screen "Screen_Doseerwals" 800x480, template "Popup_Parameters_Manual"
   on GenerateScreen: SetBit("HMI_ManualControl")
   on ClearScreen: ResetBit("HMI_ManualControl")
   TextField "Text field_1" at 624,181 size 48x23; Text 'Ready'
      Visibility <- "Drive 3 Ready"
   TextField "Text field_5" at 628,181 size 74x23; Text 'Not ready'
      Visibility <- "Drive 3 Ready"
   TextField "Template_Text field_1" at 423,141 size 182x23; Text 'Walzen - Parameters'
   TextField "Text field_3" at 10,228 size 192x23; Text 'Handbediening Walzen'
   TextField "Text field_8" at 85,262 size 42x23; Text 'Rust'
      Visibility <- "Drive 3 RUN FWD"
   TextField "Text field_9" at 103,262 size 111x23; Text 'Wals running'
      Visibility <- "Drive 3 RUN FWD"
   TextField "Text field_4" at 433,180 size 105x23; Text 'Drive Status'
   TextField "Text field_6" at 433,354 size 165x23; Text 'Reference Position:'
   IOField "StartMotorTimer" at 626,350 size 96x32; FormatPattern 9999
      ProcessValue <- "PositionManagement_Axis 3_Values_Reference Position"
   TextField "Text field_12" at 433,395 size 113x23; Text 'Rest Position'
   IOField "I/O field_2" at 625,392 size 96x32; FormatPattern 99.9999
      ProcessValue <- "PositionManagement_Axis 3_Values_Rest Position"
   Button "Button_5" at 16,389 size 111x66; TextOff '++'
      Appearance <- "Drive_3_Manual"
      on Press: SetBit("Manual Jog Fwd")
      on Release: ResetBit("Manual Jog Fwd")
   Button "Button_6" at 152,388 size 111x66; TextOff '--'
      on Release: ResetBit("Manual Jog Rev")
      on Press: SetBit("Manual Jog Rev")
   Circle "Circle_1" at 626,206 size 20x20
      Appearance <- "Voorverdeelwals staat in positie"
   Group "Group_DriveStatus" at 624,181 size 78x23
   GraphicView "Graphic view_1" at 210,135 size 172x116; Picture "MotoriconArrowLeftRight"
   Circle "Circle_2" at 221,181 size 20x20
      Appearance <- "Drive 3 REV"
   Circle "Circle_3" at 344,181 size 20x20
      Appearance <- "Drive 3 RUN FWD"
   Circle "Circle_4" at 264,229 size 16x16
      Appearance <- "Drive 3 Rapid Stop"
   TextField "Text field_2" at 210,225 size 53x23; Text 'Brake'
   TextField "Text field_10" at 13,314 size 144x23; Text 'Current Position:'
   IOField "I/O field_1" at 160,307 size 140x35; FormatPattern 9999.9999
      ProcessValue <- "PositionManagement_Data_Actual_Axis1_Position"
   TextField "Text field_11" at 433,206 size 148x23; Text 'Reference Sensor'
   TextField "Text field_13" at 433,235 size 163x23; Text 'Pulsfactor Encoder:'
   IOField "I/O field_3" at 626,229 size 96x32; FormatPattern 999.99
      ProcessValue <- "PositionManagement_Axis 3_Values_Pulsfactor"
   TextField "Text field_14" at 13,347 size 144x23; Text 'Desired Position:'
   IOField "I/O field_4" at 160,343 size 140x35; FormatPattern 999.9
      ProcessValue <- "PositionManagement_Demo_Pos_Desired_Pos"
   Button "Button_7" at 314,348 size 45x26; TextOff 'Go'
      on Press: SetBit("PositionManagement_Demo_Pos_Start")
      on Release: ResetBit("PositionManagement_Demo_Pos_Start")
   TextField "Text field_15" at 313,310 size 59x22; Text 'Degrees'
   TextField "Text field_16" at 434,275 size 101x23; Text 'Axis Speed:'
   IOField "I/O field_5" at 626,269 size 96x32; FormatPattern 99
      ProcessValue <- "PositionManagement_Axis 3_Values_Axis_Speed"
   TextField "Text field_17" at 434,314 size 163x23; Text 'Position Tolerance:'
   IOField "I/O field_6" at 626,308 size 96x32; FormatPattern 9.99
      ProcessValue <- "PositionManagement_Axis 3_Values_Position Offset"
   TextField "Text field_18" at 726,354 size 59x22; Text 'Degrees'
   TextField "Text field_19" at 727,315 size 59x22; Text 'Degrees'
   TextField "Text field_20" at 729,274 size 20x22; Text '%'
   TextField "Text field_21" at 731,234 size 41x22; Text 'Steps'
   TextField "Text field_22" at 728,396 size 59x22; Text 'Degrees'
   TextField "Text field_7" at 433,431 size 92x23; Text 'Raw Value'
   IOField "I/O field_7" at 625,428 size 96x32; FormatPattern 999999
      ProcessValue <- "Counter2_IW102"
   TextField "Text field_23" at 728,432 size 45x22; Text 'Pulses'
   Button "Button_1" at 16,149 size 126x32; TextOff 'Start Ref Run'
      on Release: ResetBit("PositionManagement_Axis 3_Commands_Start Ref Run")
      on Press: SetBit("PositionManagement_Axis 3_Commands_Start Ref Run")
      Appearance <- "Drive_3_Manual"

screen "Screen_Afdichting" 800x480, template "Popup_Parameters_Manual"
   on GenerateScreen: SetBit("HMI_ManualControl")
   on ClearScreen: ResetBit("HMI_ManualControl")
   TextField "Text field_2" at 10,228 size 290x23; Text 'Handbediening Afdichtingssysteem'
   TextField "Text field_8" at 85,262 size 42x23; Text 'Rust'
      Visibility <- "Valve 1"
   TextField "Text field_9" at 103,262 size 120x23; Text 'Valve opening'
      Visibility <- "Valve 1"
   TextField "Text field_6" at 477,376 size 247x23; Text 'Currently no parameters here'
   TextField "Template_Text field_1" at 430,142 size 205x23; Text 'Afdichting - Parameters'
   TextField "Template_Text field_2" at 12,307 size 232x23; Text 'Afdichting - Handbediening'
   Button "Button_1" at 25,340 size 110x70; TextOff 'Cilinder uit'
      on Click: SetBit("Valve_1_Manual")
      Appearance <- "Valve_1_Manual"
   Button "Button_2" at 152,340 size 110x70; TextOff 'Cilinder in'
      on Click: ResetBit("Valve_1_Manual")
   Group "Enable_Module_2" at 278,358 size 99x32; TextList "Enable / Disable List"; PictureList "Enable_Graphic"
   Group "Group" at 533,189 size 143x74; Picture "Pneumatic 5_2 valve"
   GraphicView "Graphic view_1" at 533,199 size 143x64; Picture "Pneumatic 5_2 valve"
   Circle "Circle_1" at 536,189 size 20x20
      Appearance <- "Valve 1"
   SymbolicIOField "Symbolic I/O field_3" at 311,358 size 66x32; TextOn '1'; TextOff '0'; TextList "Enable / Disable List"
      ProcessValue <- "PLCMemory_Disable_Modules_Disable_Afsluiter"
   GraphicIOField "Graphic I/O field_3" at 278,358 size 32x32; PictureList "Enable_Graphic"
      on Deactivate: ResetBit("PLCMemory_Disable_Modules_Disable_Aandruk1")
      on Activate: SetBit("PLCMemory_Disable_Modules_Disable_Aandruk1")
      ProcessValue <- "PLCMemory_Disable_Modules_Disable_Afsluiter"

screen "Screen_Settings" 800x480, template "Popup_Parameters_Manual"
   TextField "Text field_1" at 7,129 size 141x23; Text 'General Settings'
   Button "Button_7" at 487,6 size 96x65; TextOff 'Home'
      on Click: ActivateScreen("Screen_Handbediening", 0)
   TextField "Text field_12" at 420,218 size 131x23; Text 'Wals Slip Time:'
   IOField "Wals_Slip_Time" at 656,213 size 96x32; FormatPattern 9999
      ProcessValue <- "PLCMemory_WalsCheck_Time"
   TextField "Text field_13" at 420,255 size 174x23; Text 'Magazijn leeg delay:'
   IOField "I/O field_2" at 656,251 size 96x32; FormatPattern 99999
      ProcessValue <- "PLCMemory_Magazijn_Sensor_Delay"
   TextField "Template_Text field_1" at 420,154 size 186x23; Text 'General - Parameters'
   Button "Button_5" at 16,189 size 333x55; TextOff 'Manual Start'
      on Click: SetBit("RUN_Manual")
   Button "Button_6" at 15,255 size 333x55; TextOff 'Manual Stop'
      on Click: ResetBit("RUN_Manual")
   TextField "Text field_3" at 11,156 size 371x23; Text 'DO NOT USE THIS BUTTONS! IT IS DANGEROUS!'
   IOField "I/O field_1" at 656,173 size 96x32; FormatPattern 9999
      ProcessValue <- "PLCMemory_Safety_Delay"
   TextField "Text field_2" at 421,177 size 137x23; Text 'Safety on delay:'
   Button "Button_9" at 23,420 size 122x32; TextOff 'Close RT'
      on Click: StopRuntime(0)
   Button "Button_10" at 156,420 size 122x32; TextOff 'Alarms / LOG'
      on Click: ActivateScreen("AlarmWindow", 0)
   TextField "Text field_4" at 16,325 size 118x23; Text 'Invert Safety:'
   TextField "Text field_5" at 16,362 size 168x23; Text 'Invert Notensensor:'
   SymbolicIOField "Symbolic I/O field_1" at 253,317 size 96x32; TextOff '0'; TextOn '1'; TextList "List_Deactivate_Module"
      ProcessValue <- "Safety_Override"
   SymbolicIOField "Symbolic I/O field_2" at 253,353 size 96x32; TextOn '1'; TextOff '0'; TextList "List_Deactivate_Module"
      ProcessValue <- "Invert_Trechter_Sensor"
   TextField "Text field_8" at 420,295 size 174x23; Text 'Product Check Time:'
   IOField "ProductCheckTime" at 656,291 size 96x32; FormatPattern 99999
      ProcessValue <- "PLCMemory_ProductCheck_Time"
   IOField "I/O field_3" at 658,403 size 96x32; FormatPattern 999999
      ProcessValue <- "PLCMemory_TD_Products_Counter"
   TextField "Text field_6" at 422,407 size 229x23; Text 'Aantal producten gedraaid:'
   Button "Button_11" at 659,440 size 122x32; TextOff 'Reset teller'
      on Press: SetBit("ResetTotalProducts")
      on Release: ResetBit("ResetTotalProducts")
   TextField "Text field_11" at 754,176 size 25x22; Text 'ms'
   TextField "Text field_7" at 754,216 size 25x22; Text 'ms'
   TextField "Text field_9" at 754,253 size 25x22; Text 'ms'
   TextField "Text field_10" at 754,293 size 25x22; Text 'ms'
   TextField "Text field_14" at 421,334 size 169x23; Text 'BlowOff Cycle Time:'
   IOField "ProductCheckTime_1" at 657,330 size 96x32; FormatPattern 99999
      ProcessValue <- "PLCMemory_Offset_Timers_BlowOff_CycleTime"
   TextField "Text field_15" at 755,332 size 25x22; Text 'ms'
   TextField "Text field_16" at 422,372 size 170x23; Text 'BlowOff Pulse Time:'
   IOField "ProductCheckTime_2" at 658,367 size 96x32; FormatPattern 99999
      ProcessValue <- "PLCMemory_Offset_Timers_Blow_Off_PulseTime"
   TextField "Text field_17" at 756,369 size 25x22; Text 'ms'
   Softkey "Softkey_F1" at 0,0 size 0x0
      on KeyDown: function_ee5b8808("Button_7")
      on KeyUp: function_f101fd67("Button_7")

Template "Popup_Parameters" 800x480
   Rectangle "Rectangle_1" at 0,33 size 799x45
      Visibility <- "Alarm_Product_Not_Position"
   TextField "Text field_2" at 99,41 size 644x29; Text 'Aanvoer - Producten komen niet op positie, controleer sensor'
      Visibility <- "Alarm_Product_Not_Position"
   GraphicView "Graphic view_1" at 8,39 size 37x35; Picture "Graphic_30"
      Visibility <- "Alarm_Product_Not_Position"
   Group "ProductNotPositionError_1" at 0,33 size 799x45; Picture "Graphic_30"
   Group "WalsNotPositionError_1" at 0,23 size 799x45; Picture "Graphic_30"
   Group "MagazineEmptyError_1" at 0,11 size 799x45; Picture "Graphic_30"
   Group "ESB_Active_Message_2" at 0,4 size 799x45; Picture "Graphic_31"
   Group "ESB_Active_Message_1" at 1,0 size 799x45; Picture "Graphic_31"
   Rectangle "Rectangle_2" at 0,23 size 799x45
      Visibility <- "Alarm_Axis_Not_Position"
   TextField "Text field_3" at 196,31 size 395x29; Text 'Wals - As komt niet op positie of slipt'
      Visibility <- "Alarm_Axis_Not_Position"
   GraphicView "Graphic view_2" at 8,29 size 37x35; Picture "Graphic_30"
      Visibility <- "Alarm_Axis_Not_Position"
   Rectangle "Rectangle_7" at 0,11 size 799x45
      Visibility <- "Trechter_Bijvullen_Signaal"
   TextField "Text field_4" at 53,19 size 705x29; Text 'Notenmagazijn leeg - Let op, noten bijvullen om te kunnen starten!'
      Visibility <- "Trechter_Bijvullen_Signaal"
   GraphicView "Graphic view_8" at 8,17 size 37x35; Picture "Graphic_30"
      Visibility <- "Trechter_Bijvullen_Signaal"
   Rectangle "Rectangle_8" at 1,0 size 799x45
      Visibility <- "ESB_Safety_Alarm"
   GraphicView "Graphic view_9" at 10,6 size 37x35; Picture "Graphic_31"
      Visibility <- "ESB_Safety_Alarm"
   TextField "Text field_5" at 80,8 size 648x29; Text 'NOODSTOP INGEDRUKT - Ontgrendel Noodstop en druk reset'
      Visibility <- "ESB_Safety_Alarm"
   GraphicView "Graphic view_10" at 753,7 size 37x35; Picture "Graphic_31"
      Visibility <- "ESB_Safety_Alarm"
   Rectangle "Rectangle_3" at 0,4 size 799x45
      Visibility <- "Door_Safety_Alarm"
   GraphicView "Graphic view_3" at 9,10 size 37x35; Picture "Graphic_31"
      Visibility <- "Door_Safety_Alarm"
   TextField "Text field_1" at 174,12 size 511x29; Text 'DEUR(EN) OPEN - Sluit alle deuren en druk reset'
      Visibility <- "Door_Safety_Alarm"
   GraphicView "Graphic view_4" at 752,11 size 37x35; Picture "Graphic_31"
      Visibility <- "Door_Safety_Alarm"
   Group "Message_Group_General" at 0,0 size 800x78; Picture "Graphic_30"

Template "Popup_Parameters_Manual" 800x480
   Rectangle "Rectangle_1" at 0,106 size 799x45
      Visibility <- "Alarm_Product_Not_Position"
   TextField "Text field_2" at 99,114 size 644x29; Text 'Aanvoer - Producten komen niet op positie, controleer sensor'
      Visibility <- "Alarm_Product_Not_Position"
   GraphicView "Graphic view_1" at 8,112 size 37x35; Picture "Graphic_30"
      Visibility <- "Alarm_Product_Not_Position"
   Group "ProductNotPositionError_1" at 0,106 size 799x45; Picture "Graphic_30"
   Group "WalsNotPositionError_1" at 0,96 size 799x45; Picture "Graphic_30"
   Group "MagazineEmptyError_1" at 0,84 size 799x45; Picture "Graphic_30"
   Group "ESB_Active_Message_2" at 0,77 size 799x45; Picture "Graphic_31"
   Group "ESB_Active_Message_1" at 1,73 size 799x45; Picture "Graphic_31"
   Rectangle "Rectangle_2" at 0,96 size 799x45
      Visibility <- "Alarm_Axis_Not_Position"
   TextField "Text field_3" at 196,104 size 395x29; Text 'Wals - As komt niet op positie of slipt'
      Visibility <- "Alarm_Axis_Not_Position"
   GraphicView "Graphic view_2" at 8,102 size 37x35; Picture "Graphic_30"
      Visibility <- "Alarm_Axis_Not_Position"
   Rectangle "Rectangle_7" at 0,84 size 799x45
      Visibility <- "Trechter_Bijvullen_Signaal"
   TextField "Text field_4" at 53,92 size 705x29; Text 'Notenmagazijn leeg - Let op, noten bijvullen om te kunnen starten!'
      Visibility <- "Trechter_Bijvullen_Signaal"
   GraphicView "Graphic view_8" at 8,90 size 37x35; Picture "Graphic_30"
      Visibility <- "Trechter_Bijvullen_Signaal"
   Rectangle "Rectangle_3" at 0,77 size 799x45
      Visibility <- "Door_Safety_Alarm"
   GraphicView "Graphic view_3" at 9,83 size 37x35; Picture "Graphic_31"
      Visibility <- "Door_Safety_Alarm"
   TextField "Text field_1" at 174,85 size 511x29; Text 'DEUR(EN) OPEN - Sluit alle deuren en druk reset'
      Visibility <- "Door_Safety_Alarm"
   GraphicView "Graphic view_4" at 752,84 size 37x35; Picture "Graphic_31"
      Visibility <- "Door_Safety_Alarm"
   Rectangle "Rectangle_8" at 1,73 size 799x45
      Visibility <- "ESB_Safety_Alarm"
   GraphicView "Graphic view_9" at 10,79 size 37x35; Picture "Graphic_31"
      Visibility <- "ESB_Safety_Alarm"
   TextField "Text field_5" at 80,81 size 648x29; Text 'NOODSTOP INGEDRUKT - Ontgrendel Noodstop en druk reset'
      Visibility <- "ESB_Safety_Alarm"
   GraphicView "Graphic view_10" at 753,80 size 37x35; Picture "Graphic_31"
      Visibility <- "ESB_Safety_Alarm"
   TextField "Text field_7" at 14,261 size 70x23; Text 'Sturing:'
   Button "Button_3" at 693,5 size 100x65; TextOff 'Logoff'
      on Click: function_f23ef4c9()
   Button "Button_4" at 585,5 size 100x65; TextOff 'Back'
      on Click: function_efd93a16()
   Group "Message_Group_Manual" at 0,73 size 800x78; Picture "Graphic_30"

screen "Screen_Automatiek" 800x480, template "Popup_Parameters"
   Softkey "Softkey_F8" at 0,0 size 0x0
      on KeyDown: function_ee5b8808("Button_3")
      on KeyUp: function_f101fd67("Button_3")
   TextField "Text field_1" at 263,165 size 182x23; Text 'Gekozen Programma:'
   TextField "Text field_2" at 451,166 size 15x23; Text '1'
      Appearance <- "LED Programma 1"
   TextField "Text field_3" at 469,166 size 15x23; Text '2'
      Appearance <- "LED Programma 2"
   TextField "Text field_4" at 489,166 size 15x23; Text '3'
      Appearance <- "LED Programma 3"
   Button "Button_3" at 6,157 size 130x60; TextOn 'Onderweg na vorig scherm'; TextOff 'Terug'
      on Click: function_efd93a16()
   Button "Button_1" at 6,222 size 130x60; TextOn 'Onderweg na vorig scherm'; TextOff 'Instellingen'
      on Click: ActivateScreen("Screen_Settings", 0)
   TextField "Text field_5" at 26,112 size 106x23; Text 'Automatiek'
   TextField "Text field_6" at 608,165 size 144x23; Text 'Product Interval:'
   IOField "I/O field_1" at 610,189 size 96x32; FormatPattern 99999
      ProcessValue <- "PLCMemory_ProductIntervalTime"
   TextField "Text field_11" at 710,197 size 68x22; Text 'Seconden'
   TextField "Text field_7" at 292,263 size 179x23; Text 'Aanvoerband Gestart'
      Appearance <- "Drive 1 Ready"
      Visibility <- "Drive 1 RUN FWD"
   TextField "Text field_8" at 299,224 size 160x23; Text 'Koek gedetecteerd'
      Visibility <- "Sensor_op_band_memory"
   TextField "Text field_9" at 290,374 size 178x23; Text 'Doseerwals Draaiend'
      Appearance <- "Drive 3 Ready"
      Visibility <- "PLCMemory_ProductBuffer_MoveTrigger"
   TextField "Text field_10" at 282,337 size 196x23; Text 'Aanvoer Wals Draaiend'
      Visibility <- "Drive 4 RUN FWD"
   TextField "Text field_12" at 308,300 size 146x23; Text 'Trilgoten Gestart'
      Appearance <- "Drive 2 Ready"
      Visibility <- "Drive 2 RUN FWD"
   TextField "Text field_13" at 306,189 size 166x23; Text 'Programma Started'
      Visibility <- "Systeem RUN"
   TextField "Text field_14" at 308,419 size 155x23; Text 'Programma Ended'
      Visibility <- "Systeem RUN"
   GraphicView "Graphic view_1" at 371,209 size 26x22; Picture "Graphic_32"
   GraphicView "Graphic view_2" at 371,246 size 26x22; Picture "Graphic_32"
   GraphicView "Graphic view_3" at 372,283 size 26x22; Picture "Graphic_32"
   GraphicView "Graphic view_4" at 371,320 size 26x22; Picture "Graphic_32"
   GraphicView "Graphic view_5" at 372,357 size 26x22; Picture "Graphic_32"
   GraphicView "Graphic view_6" at 372,399 size 26x22; Picture "Graphic_32"
   TextField "Text field_15" at 608,222 size 123x23; Text 'Product Buffer'
   IOField "I/O field_2" at 610,246 size 96x32; FormatPattern 999
      ProcessValue <- "PLCMemory_ProductBuffer_ProductsCount"
   TextField "Text field_16" at 710,254 size 70x22; Text 'Producten'
   TextField "Text field_17" at 608,281 size 129x23; Text 'Aandruk Buffer'
   IOField "I/O field_3" at 610,305 size 96x32; FormatPattern 99
      ProcessValue <- "PLCMemory_ProductBufferBehindWals_Product_Count"
   TextField "Text field_18" at 710,313 size 70x22; Text 'Producten'
   Button "Button_2" at 6,286 size 130x60; TextOn 'Onderweg na vorig scherm'; TextOff 'Buffer Data'
      on Click: ActivateScreen("Screen_Automatiek_BufferData", 0)

screen "Screen_Trechterwissel" 800x480, template "Popup_Parameters_Manual"
   TextField "Text field_2" at 10,228 size 324x23; Text 'Handbediening Trechter wisselsysteem'
   TextField "Text field_8" at 85,262 size 42x23; Text 'Rust'
      Visibility <- "Valve 2"
   TextField "Text field_9" at 103,262 size 120x23; Text 'Valve opening'
      Visibility <- "Valve 2"
   TextField "Template_Text field_1" at 423,142 size 241x23; Text 'Wisselsysteem - Parameters'
   TextField "Template_Text field_2" at 12,307 size 268x23; Text 'Wisselsysteem - Handbediening'
   Button "Button_1" at 17,338 size 111x32; TextOff 'Cilinder uit'
      on Click: SetBit("Valve_2_Manual")
      Appearance <- "Valve_2_Manual"
   Button "Button_2" at 152,338 size 111x32; TextOff 'Cilinder in'
      on Click: ResetBit("Valve_2_Manual")
   GraphicView "Graphic view_1" at 533,197 size 143x64; Picture "Pneumatic 5_2 valve"
   Circle "Circle_1" at 536,187 size 20x20
      Appearance <- "Valve 2"
   TextField "Text field_13" at 12,381 size 173x23; Text 'Reedcontact Cilinder in:'
   Circle "Circle_2" at 198,384 size 20x20
      Appearance <- "Cilinder Trechterwissel in"
   TextField "Text field_1" at 12,407 size 178x23; Text 'Reedcontact Cilinder uit:'
   Circle "Circle_3" at 198,410 size 20x20
      Appearance <- "Cilinder Trechterwissel uit"
   TextField "Text field_12" at 429,337 size 181x23; Text 'Delay Wisselsysteem:'
   IOField "I/O field_2" at 620,334 size 96x32; FormatPattern 9999

screen "Screen_Aandrukken" 800x480, template "Popup_Parameters_Manual"
   on ClearScreen: ResetBit("HMI_ManualControl")
   on GenerateScreen: SetBit("HMI_ManualControl")
   TextField "Text field_2" at 10,228 size 268x23; Text 'Handbediening Aandruksysteem'
   TextField "Text field_8" at 85,262 size 42x23; Text 'Rust'
      Visibility <- "Valve 3"
   TextField "Text field_9" at 103,262 size 120x23; Text 'Valve opening'
      Visibility <- "Valve 3"
   Button "Button_1" at 428,144 size 110x70; TextOff 'Cilinder 1 uit'
      on Click: SetBit("Valve_3_Manual")
      Appearance <- "Valve_3_Manual"
   Button "Button_2" at 555,144 size 110x70; TextOff 'Cilinder 1 in'
      on Click: ResetBit("Valve_3_Manual")
   Button "Button_5" at 428,241 size 110x70; TextOff 'Cilinder 2 uit'
      on Click: SetBit("Valve_4_Manual")
      Appearance <- "Valve_4_Manual"
   Button "Button_6" at 555,241 size 110x70; TextOff 'Cilinder 2 in'
      on Click: ResetBit("Valve_4_Manual")
   Button "Button_7" at 428,338 size 110x70; TextOff 'Cilinder 3 uit'
      on Click: SetBit("Valve_5_Manual")
      Appearance <- "Valve_5_Manual"
   Button "Button_8" at 555,338 size 110x70; TextOff 'Cilinder 3 in'
      on Click: ResetBit("Valve_5_Manual")
   Button "Button_10" at 24,402 size 150x55; TextOff 'Alle cilinders uit'
      on Click: SetBit("Valve_3_Manual"); SetBit("Valve_4_Manual"); SetBit("Valve_5_Manual")
      Appearance <- "Valve_3_Manual"
   Button "Button_11" at 218,402 size 150x55; TextOff 'Alle cilinders in'
      on Click: ResetBit("Valve_3_Manual"); ResetBit("Valve_4_Manual"); ResetBit("Valve_5_Manual")
   Group "Group" at 15,301 size 207x87; Picture "Pneumatic 5_2 valve"
   Button "Button_3" at 127,351 size 150x45; TextOff 'Blaaspuls aan'
      Appearance <- "Valve_3_Manual"
      on Release: ResetBit("Valve_2_Manual")
      on Press: SetBit("Valve_2_Manual")
   Group "Enable_Module" at 684,163 size 99x32; TextList "Enable / Disable List"; PictureList "Enable_Graphic"
   Group "Enable_Module_1" at 683,264 size 99x32; TextList "Enable / Disable List"; PictureList "Enable_Graphic"
   Group "Enable_Module_2" at 684,357 size 99x32; PictureList "Enable_Graphic"; TextList "Enable / Disable List"
   Group "Enable_Module_3" at 279,356 size 99x32; TextList "Enable / Disable List"; PictureList "Enable_Graphic"
   GraphicView "Graphic view_1" at 16,307 size 95x37; Picture "Pneumatic 5_2 valve"
   GraphicView "Graphic view_2" at 127,307 size 95x37; Picture "Pneumatic 5_2 valve"
   Circle "Circle_2" at 130,301 size 12x12
      Appearance <- "Valve 5"
   Circle "Circle_1" at 19,301 size 12x12
      Appearance <- "Valve 3"
   GraphicView "Graphic view_3" at 15,351 size 95x37; Picture "Pneumatic 5_2 valve"
   Circle "Circle_3" at 18,345 size 12x12
      Appearance <- "Valve 4"
   TextField "Text field_1" at 64,304 size 15x23; Text '1'
   TextField "Text field_3" at 64,348 size 15x23; Text '2'
   TextField "Text field_4" at 176,305 size 15x23; Text '3'
   SymbolicIOField "Symbolic I/O field_2" at 717,163 size 66x32; TextOn '1'; TextOff '0'; TextList "Enable / Disable List"
      ProcessValue <- "PLCMemory_Disable_Modules_Disable_Aandruk1"
   GraphicIOField "Graphic I/O field_1" at 684,163 size 32x32; PictureList "Enable_Graphic"
      ProcessValue <- "PLCMemory_Disable_Modules_Disable_Aandruk1"
      on Activate: SetBit("PLCMemory_Disable_Modules_Disable_Aandruk1")
      on Deactivate: ResetBit("PLCMemory_Disable_Modules_Disable_Aandruk1")
   SymbolicIOField "Symbolic I/O field_1" at 716,264 size 66x32; TextOn '1'; TextOff '0'; TextList "Enable / Disable List"
      ProcessValue <- "PLCMemory_Disable_Modules_Disable_Aandruk2"
   GraphicIOField "Graphic I/O field_2" at 683,264 size 32x32; PictureList "Enable_Graphic"
      on Deactivate: ResetBit("PLCMemory_Disable_Modules_Disable_Aandruk1")
      on Activate: SetBit("PLCMemory_Disable_Modules_Disable_Aandruk1")
      ProcessValue <- "PLCMemory_Disable_Modules_Disable_Aandruk2"
   SymbolicIOField "Symbolic I/O field_3" at 717,357 size 66x32; TextOn '1'; TextOff '0'; TextList "Enable / Disable List"
      ProcessValue <- "PLCMemory_Disable_Modules_Disable_Aandruk3"
   GraphicIOField "Graphic I/O field_3" at 684,357 size 32x32; PictureList "Enable_Graphic"
      on Deactivate: ResetBit("PLCMemory_Disable_Modules_Disable_Aandruk1")
      on Activate: SetBit("PLCMemory_Disable_Modules_Disable_Aandruk1")
      ProcessValue <- "PLCMemory_Disable_Modules_Disable_Aandruk3"
   SymbolicIOField "Symbolic I/O field_4" at 312,356 size 66x32; TextOn '1'; TextOff '0'; TextList "Enable / Disable List"
      ProcessValue <- "PLCMemory_Disable_Modules_Disable_Blaaspuls"
   GraphicIOField "Graphic I/O field_4" at 279,356 size 32x32; PictureList "Enable_Graphic"
      on Deactivate: ResetBit("PLCMemory_Disable_Modules_Disable_Aandruk1")
      on Activate: SetBit("PLCMemory_Disable_Modules_Disable_Aandruk1")
      ProcessValue <- "PLCMemory_Disable_Modules_Disable_Blaaspuls"

screen "Screen_RetourBand" 800x480, template "Popup_Parameters_Manual"
   on GenerateScreen: SetBit("HMI_ManualControl")
   on ClearScreen: ResetBit("HMI_ManualControl")
   TextField "Text field_1" at 8,220 size 255x23; Text 'Handbediening Retoursysteem'
   TextField "Text field_8" at 85,261 size 42x23; Text 'Rust'
      Visibility <- "Drive 5 Ready"
   TextField "Text field_9" at 103,261 size 113x23; Text 'Band running'
      Visibility <- "Drive 5 Ready"
   TextField "Text field_3" at 426,174 size 105x23; Text 'Drive Status'
   TextField "Text field_2" at 426,228 size 153x23; Text 'Start Timer motor'
   IOField "StartMotorTimer" at 584,224 size 96x32; FormatPattern 9999
   TextField "Text field_6" at 426,262 size 149x23; Text 'Stop Timer motor'
   IOField "I/O field_2" at 584,259 size 96x32; FormatPattern 9999
   TextField "Template_Text field_1" at 426,140 size 218x23; Text 'Retourband - Parameters'
   Button "Button_1" at 25,306 size 135x70; TextOff 'Start FWD'
      on Click: SetBit("Drive_5_Manual")
      Appearance <- "Drive_1_Manual"
   Button "Button_2" at 205,306 size 135x70; TextOff 'Stop FWD'
      on Click: ResetBit("Drive_5_Manual")
      on Release: ResetBit("Stop_drive_1")
      on Press: SetBit("Stop_drive_1")
   Button "Button_5" at 25,390 size 135x70; TextOff 'Start Rev'
      on Click: SetBit("Drive 5 REV")
      Appearance <- "Drive 5 REV"
   Button "Button_6" at 205,390 size 135x70; TextOff 'Stop Rev'
      on Click: ResetBit("Drive 5 REV")
   Group "Group" at 582,174 size 77x23
   GraphicView "Graphic view_1" at 272,133 size 135x113; Picture "MotoriconArrowLeftRight"
   Circle "Circle_1" at 277,176 size 20x20
      Appearance <- "Drive 5 REV"
   Circle "Circle_2" at 377,176 size 20x20
      Appearance <- "Drive 5 RUN FWD"
   Circle "Circle_3" at 585,199 size 20x20
      Appearance <- "Drive 5 Rapid Stop"
   TextField "Text field_12" at 426,200 size 101x23; Text 'Drive Brake'
   TextField "Text field_13" at 688,228 size 25x22; Text 'ms'
   TextField "Text field_14" at 688,265 size 25x22; Text 'ms'
   Group "Enable_Module" at 584,298 size 96x32; TextList "Enable / Disable List"; PictureList "Enable_Graphic"
   TextField "Text field_7" at 426,302 size 108x23; Text 'Enable Drive'
   TextField "Text field_5" at 582,174 size 48x23; Text 'Ready'
      Visibility <- "Drive 5 Ready"
   TextField "Text field_4" at 585,174 size 74x23; Text 'Not ready'
      Visibility <- "Drive 5 Ready"
   SymbolicIOField "Symbolic I/O field_2" at 616,298 size 64x32; TextOn '1'; TextOff '0'; TextList "Enable / Disable List"
      ProcessValue <- "PLCMemory_Disable_Modules_Disable_Retourband"
   GraphicIOField "Graphic I/O field_1" at 584,298 size 31x32; PictureList "Enable_Graphic"
      on Deactivate: ResetBit("PLCMemory_Disable_Modules_Disable_Aandruk1")
      on Activate: SetBit("PLCMemory_Disable_Modules_Disable_Aandruk1")
      ProcessValue <- "PLCMemory_Disable_Modules_Disable_Retourband"

screen "Screen_Safety_I/O" 800x480, template "Popup_Parameters"
   TextField "Text field_1" at 185,162 size 145x23; Text 'Noodstop Status:'
   Button "Button_4" at 6,157 size 130x60; TextOn 'Onderweg na vorig scherm'; TextOff 'Terug'
      on Click: function_efd93a16()
   Button "Button_5" at 6,221 size 130x60; TextOn 'Onderweg na vorig scherm'; TextOff 'Instellingen'
      on Click: ActivateScreen("Screen_Settings", 0)
   TextField "Text field_2" at 26,112 size 173x23; Text 'Safety In en Outputs'
   TextField "Text field_6" at 185,221 size 122x23; Text 'Deur 1 Status:'
   TextField "Text field_3" at 185,252 size 122x23; Text 'Deur 2 Status:'
   TextField "Text field_4" at 185,281 size 175x23; Text 'Safety Relais Status:'
   TextField "Text field_7" at 185,194 size 115x23; Text 'Reset Status:'
   Circle "Circle_1" at 394,164 size 21x21
      Appearance <- "ESB Oke"
   Circle "Circle_2" at 396,221 size 21x21
      Appearance <- "Door 1 NC contact"
   Circle "Circle_3" at 396,252 size 21x21
      Appearance <- "Door 2 NC contact"
   Circle "Circle_4" at 396,193 size 21x21
      Appearance <- "Reset Active"
   Circle "Circle_5" at 397,284 size 21x21
      Appearance <- "Safety Relais"
   TextField "Text field_8" at 185,309 size 136x23; Text 'Safety override:'
   TextField "Text field_9" at 394,311 size 56x23; Text 'Active'
      Visibility <- "Safety_Override"
   TextField "Text field_10" at 397,311 size 90x23; Text 'Not Active'
      Visibility <- "Safety_Override"

screen "AlarmWindow" 800x480, template "Popup_Parameters"
   AlarmView "Alarm view_1" at 5,119 size 782x352
   Button "Button_1" at 690,82 size 96x32; TextOff 'Sluiten'
      on Click: function_efd93a16()
   Button "Button_2" at 532,82 size 147x32; TextOff 'Reset Storingen'
      on Release: function_a9b64e44("Clear_Error", 0); function_a9b64e44("Clear_Error", 1); function_a9b64e44("Clear_Error", 2); function_a9b64e44("Clear_Error", 3); function_a9b64e44("Clear_Error", 4); function_a9b64e44("Clear_Error", 5); function_a9b64e44("Clear_Error", 6)
      on Press: function_b3f726e6("Clear_Error", 0); function_b3f726e6("Clear_Error", 1); function_b3f726e6("Clear_Error", 2); function_b3f726e6("Clear_Error", 3); function_b3f726e6("Clear_Error", 4); function_b3f726e6("Clear_Error", 5); function_b3f726e6("Clear_Error", 6)
      on Click: function_dcc94856(-1); function_e14cd482(0)

screen "Screen_Infeed" 800x480, template "Popup_Parameters"
   on ClearScreen: ResetBit("HMI_ManualControl")
   on GenerateScreen: SetBit("HMI_ManualControl")
   Button "Button_2" at 47,158 size 130x60; TextOn 'Onderweg na vorig scherm'; TextOff 'Terug'
      on Click: function_efd93a16()
   TextField "Text field_10" at 62,125 size 124x23; Text 'Invoer Koeken'
   Button "Button_4" at 263,155 size 184x60; TextOn 'Onderweg na vorig scherm'; TextOff 'Aanvoer Wals Noten'
      on Click: ActivateScreen("Screen_AanvoerWals", 0)
   Button "Button_5" at 573,158 size 130x60; TextOn 'Onderweg na vorig scherm'; TextOff 'Invoerband'
      on Click: ActivateScreen("Screen_Band", 0)
   GraphicView "Graphic view_1" at 314,86 size 95x61; Picture "MotoriconArrowLeftRight"
   GraphicView "Graphic view_2" at 591,86 size 95x61; Picture "MotoriconArrowLeftRight"

screen "Screen_AanvoerWals" 800x480, template "Popup_Parameters_Manual"
   on GenerateScreen: SetBit("HMI_ManualControl")
   on ClearScreen: ResetBit("HMI_ManualControl")
   TextField "Text field_8" at 85,262 size 42x23; Text 'Rust'
      Visibility <- "Drive 4 Ready"
   TextField "Text field_9" at 103,262 size 111x23; Text 'Wals running'
      Visibility <- "Drive 4 Ready"
   TextField "Text field_3" at 423,183 size 105x23; Text 'Drive Status'
   TextField "Text field_2" at 422,238 size 147x23; Text 'Speed as Drive 1:'
   TextField "Template_Text field_1" at 423,141 size 227x23; Text 'Aanvoerwals - Parameters'
   Button "Button_1" at 25,306 size 135x70; TextOff 'Start FWD'
      on Click: SetBit("Drive_4_Manual")
      Appearance <- "Drive_4_Manual"
   Button "Button_2" at 205,306 size 135x70; TextOff 'Stop FWD'
      on Click: ResetBit("Drive_4_Manual")
      on Release: ResetBit("Stop_drive_1")
      on Press: SetBit("Stop_drive_1")
   Button "Button_5" at 25,390 size 135x70; TextOff 'Start Rev'
      on Click: SetBit("Drive 4 REV")
      Appearance <- "Drive 4 REV"
   Button "Button_6" at 205,390 size 135x70; TextOff 'Stop Rev'
      on Click: ResetBit("Drive 4 REV")
   Group "Group" at 579,183 size 77x23
   GraphicView "Graphic view_1" at 227,133 size 179x113; Picture "MotoriconArrowLeftRight"
   Circle "Circle_1" at 243,176 size 20x20
      Appearance <- "Drive 4 REV"
   Circle "Circle_2" at 369,176 size 20x20
      Appearance <- "Drive 4 RUN FWD"
   Circle "Circle_3" at 582,208 size 20x20
      Appearance <- "Drive 4 Rapid Stop"
   TextField "Text field_12" at 423,209 size 101x23; Text 'Drive Brake'
   SymbolicIOField "Symbolic I/O field_1" at 581,233 size 184x32; TextOn '1'; TextOff '0'; TextList "SpeedSettings"; HelpText 'Choose of the speed of Drive 4 is synchronized with Drive 1.'
      ProcessValue <- "PLCMemory_SpeedSettingsTakeover"
   TextField "Text field_13" at 422,351 size 153x23; Text 'Start Timer motor'
   IOField "I/O field_3" at 580,348 size 96x32; FormatPattern 9999
      ProcessValue <- "PLCMemory_Overname_Start_Offset"
   TextField "Text field_15" at 684,354 size 25x22; Text 'ms'
   TextField "Text field_6" at 424,316 size 125x23; Text 'Speed settings'
   SymbolicIOField "Symbolic I/O field_2" at 581,311 size 184x32; TextOn '1'; TextOff '0'; TextList "SpeedSettingOvername"; HelpText 'Choose the speed settings for Drive 4 when its not linked to Drive 1.'
      ProcessValue <- "PLCMemory_SpeedSettingOvername"
   TextField "Text field_14" at 424,277 size 153x23; Text 'Timing as Drive 1:'
   SymbolicIOField "Symbolic I/O field_3" at 583,272 size 184x32; TextOn '1'; TextOff '0'; TextList "SpeedSettings"; HelpText 'Choose of the Start/Stop timing of Drive 4 is synchronized with Drive 1.'
      ProcessValue <- "PLCMemory_TimingSettingOvername"
   TextField "Text field_16" at 422,386 size 149x23; Text 'Stop Timer motor'
   IOField "I/O field_2" at 580,383 size 96x32; FormatPattern 9999
      ProcessValue <- "PLCMemory_Overname_Stop_Offset"
   TextField "Text field_17" at 684,389 size 25x22; Text 'ms'
   TextField "Text field_1" at 8,220 size 244x23; Text 'Handbediening Aanvoer Wals'
   TextField "Text field_5" at 579,183 size 48x23; Text 'Ready'
      Visibility <- "Drive 4 Ready"
   TextField "Text field_4" at 582,183 size 74x23; Text 'Not ready'
      Visibility <- "Drive 4 Ready"

screen "Screen_Automatiek_BufferData" 800x480, template "Popup_Parameters"
   Softkey "Softkey_F8" at 0,0 size 0x0
      on KeyUp: function_f101fd67("Button_3")
      on KeyDown: function_ee5b8808("Button_3")
   Button "Button_1" at 6,226 size 130x60; TextOn 'Onderweg na vorig scherm'; TextOff 'Enlarge Buffer Data'
      on Click: ActivateScreen("Screen_Automatiek_BufferData_Enlarge", 0)
   TextField "Text field_1" at 194,169 size 218x23; Text 'Product Detection Sensor:'
   Button "Button_3" at 6,157 size 130x60; TextOn 'Onderweg na vorig scherm'; TextOff 'Terug'
      on Click: function_efd93a16()
   TextField "Text field_5" at 26,112 size 285x23; Text 'Automatiek - Product Buffer Data'
   TextField "Text field_6" at 608,165 size 144x23; Text 'Product Interval:'
   IOField "I/O field_1" at 610,189 size 96x32; FormatPattern 99999
      ProcessValue <- "PLCMemory_ProductIntervalTime"
   TextField "Text field_11" at 710,197 size 68x22; Text 'Seconden'
   GraphicView "Graphic view_6" at 105,243 size 28x25; Picture "Graphic_32"
   TextField "Text field_15" at 608,222 size 123x23; Text 'Product Buffer'
   IOField "I/O field_2" at 610,246 size 96x32; FormatPattern 999
      ProcessValue <- "PLCMemory_ProductBuffer_ProductsCount"
   TextField "Text field_16" at 710,254 size 70x22; Text 'Producten'
   TextField "Text field_17" at 608,281 size 129x23; Text 'Aandruk Buffer'
   IOField "I/O field_3" at 610,305 size 96x32; FormatPattern 99
      ProcessValue <- "PLCMemory_ProductBufferBehindWals_Product_Count"
   TextField "Text field_18" at 710,313 size 70x22; Text 'Producten'
   IOField "I/O field_4" at 421,165 size 96x32; FormatPattern 1
      ProcessValue <- "ProductBuffer_V2_DB_SensorInput"
   TextField "Text field_2" at 194,211 size 168x23; Text 'Trigger Delay Time:'
   IOField "I/O field_5" at 420,202 size 96x32; FormatPattern 9999999
      ProcessValue <- "PLCMemory_ProductBuffer_DelayTime"
   TextField "Text field_3" at 520,205 size 68x22; Text 'Seconden'
   TextField "Text field_4" at 195,244 size 112x23; Text 'Insert Index:'
   IOField "I/O field_6" at 421,241 size 96x32; FormatPattern 99
      ProcessValue <- "PLCMemory_ProductBuffer_InsertIndex"
   TextField "Text field_7" at 195,283 size 152x23; Text 'PLC System Time:'
   IOField "I/O field_7" at 421,278 size 116x32; FormatPattern 9999999999999
      ProcessValue <- "PLCMemory_SystemTime"
   TextField "Text field_8" at 196,320 size 126x23; Text 'Motion Trigger'
   IOField "I/O field_8" at 423,316 size 96x32; FormatPattern 1
      ProcessValue <- "ProductBuffer_V2_DB_TriggerMovement"
   TextField "Text field_9" at 195,358 size 143x23; Text 'Motion Feedback'
   IOField "I/O field_9" at 422,354 size 96x32; FormatPattern 1
      ProcessValue <- "ProductBuffer_V2_DB_TriggerFeedback"

screen "Screen_Automatiek_BufferData_Enlarge" 800x480, template "Popup_Parameters"
   Softkey "Softkey_F8" at 0,0 size 0x0
      on KeyUp: function_f101fd67("Button_3")
      on KeyDown: function_ee5b8808("Button_3")
   TextField "Text field_1" at 151,97 size 108x23; Text 'StartTime 0:'
   Button "Button_3" at 6,109 size 130x60; TextOn 'Onderweg na vorig scherm'; TextOff 'Terug'
      on Click: function_efd93a16()
   TextField "Text field_5" at 47,212 size 28x202; Text 'BufferData_Enlarged'
   IOField "I/O field_4" at 266,93 size 96x32; FormatPattern 9999999999
      ProcessValue <- "ProductBuffer_V2_DB_StartTimes__0"
   TextField "Text field_2" at 151,138 size 108x23; Text 'StartTime 1:'
   IOField "I/O field_5" at 266,133 size 96x32; FormatPattern 9999999999
      ProcessValue <- "ProductBuffer_V2_DB_StartTimes__1"
   TextField "Text field_3" at 151,177 size 108x23; Text 'StartTime 2:'
   IOField "I/O field_6" at 266,172 size 96x32; FormatPattern 9999999999
      ProcessValue <- "ProductBuffer_V2_DB_StartTimes__2"
   TextField "Text field_4" at 151,216 size 108x23; Text 'StartTime 3:'
   IOField "I/O field_7" at 266,211 size 96x32; FormatPattern 9999999999
      ProcessValue <- "ProductBuffer_V2_DB_StartTimes__3"
   TextField "Text field_7" at 151,255 size 108x23; Text 'StartTime 4:'
   IOField "I/O field_8" at 266,250 size 96x32; FormatPattern 9999999999
      ProcessValue <- "ProductBuffer_V2_DB_StartTimes__4"
   TextField "Text field_8" at 151,294 size 108x23; Text 'StartTime 5:'
   IOField "I/O field_9" at 266,289 size 96x32; FormatPattern 9999999999
      ProcessValue <- "ProductBuffer_V2_DB_StartTimes__5"
   TextField "Text field_9" at 151,333 size 108x23; Text 'StartTime 6:'
   IOField "I/O field_10" at 266,328 size 96x32; FormatPattern 9999999999
      ProcessValue <- "ProductBuffer_V2_DB_StartTimes__6"
   TextField "Text field_10" at 151,373 size 108x23; Text 'StartTime 7:'
   IOField "I/O field_11" at 266,368 size 96x32; FormatPattern 9999999999
      ProcessValue <- "ProductBuffer_V2_DB_StartTimes__7"
   TextField "Text field_12" at 151,413 size 108x23; Text 'StartTime 8:'
   IOField "I/O field_12" at 266,408 size 96x32; FormatPattern 9999999999
      ProcessValue <- "ProductBuffer_V2_DB_StartTimes__8"
   TextField "Text field_13" at 151,453 size 108x23; Text 'StartTime 9:'
   IOField "I/O field_13" at 266,448 size 96x32; FormatPattern 9999999999
      ProcessValue <- "ProductBuffer_V2_DB_StartTimes__9"
   TextField "Text field_6" at 377,93 size 85x23; Text 'Actives 0:'
   IOField "I/O field_1" at 471,89 size 96x32; FormatPattern 1
      ProcessValue <- "ProductBuffer_V2_DB_Actives__0"
   TextField "Text field_11" at 377,134 size 85x23; Text 'Actives 1:'
   IOField "I/O field_2" at 471,129 size 96x32; FormatPattern 1
      ProcessValue <- "ProductBuffer_V2_DB_Actives__1"
   TextField "Text field_14" at 377,173 size 85x23; Text 'Actives 2:'
   IOField "I/O field_3" at 471,168 size 96x32; FormatPattern 1
      ProcessValue <- "ProductBuffer_V2_DB_Actives__2"
   TextField "Text field_15" at 377,212 size 85x23; Text 'Actives 3:'
   IOField "I/O field_14" at 471,207 size 96x32; FormatPattern 1
      ProcessValue <- "ProductBuffer_V2_DB_Actives__3"
   TextField "Text field_16" at 377,251 size 85x23; Text 'Actives 4:'
   IOField "I/O field_15" at 471,246 size 96x32; FormatPattern 1
      ProcessValue <- "ProductBuffer_V2_DB_Actives__4"
   TextField "Text field_17" at 377,290 size 85x23; Text 'Actives 5:'
   IOField "I/O field_16" at 471,285 size 96x32; FormatPattern 1
      ProcessValue <- "ProductBuffer_V2_DB_Actives__5"
   TextField "Text field_18" at 377,329 size 85x23; Text 'Actives 6:'
   IOField "I/O field_17" at 471,324 size 96x32; FormatPattern 1
      ProcessValue <- "ProductBuffer_V2_DB_Actives__6"
   TextField "Text field_19" at 377,369 size 85x23; Text 'Actives 7:'
   IOField "I/O field_18" at 471,364 size 96x32; FormatPattern 1
      ProcessValue <- "ProductBuffer_V2_DB_Actives__7"
   TextField "Text field_20" at 377,409 size 85x23; Text 'Actives 8:'
   IOField "I/O field_19" at 471,404 size 96x32; FormatPattern 1
      ProcessValue <- "ProductBuffer_V2_DB_Actives__8"
   TextField "Text field_21" at 377,449 size 85x23; Text 'Actives 9:'
   IOField "I/O field_20" at 471,444 size 96x32; FormatPattern 1
      ProcessValue <- "ProductBuffer_V2_DB_Actives__9"
   TextField "Text field_22" at 592,98 size 74x23; Text 'Elapsed:'
   IOField "I/O field_21" at 676,94 size 96x32; FormatPattern 9999999999
      ProcessValue <- "ProductBuffer_V2_DB_Elapsed"
   TextField "Text field_23" at 592,137 size 83x23; Text 'Prev Sen:'
   IOField "I/O field_22" at 676,133 size 96x32; FormatPattern 1
      ProcessValue <- "ProductBuffer_V2_DB_PrevSensor"
   TextField "Text field_24" at 591,178 size 76x23; Text 'Mov Act:'
   IOField "I/O field_23" at 675,174 size 96x32; FormatPattern 1
      ProcessValue <- "ProductBuffer_V2_DB_MovementActive"
   TextField "Text field_25" at 71,235 size 21x150; Text 'All Data in Milliseconds'
*)